(* Logix 5000 project; controller MV vendor 1 type 14 code 217 rev 31.11; software revision 31.00 *)

TASK _1Sec (periodic, rate 1000 ms, priority 10, watchdog 500 ms) : _1Second
TASK MainTask (continuous, watchdog 500 ms) : First_Task, MV_Common, MC_Common, Last_Task

MODULES
   Local : vendor 1 type 14 code 217 (5069 0, rev 31.11)
      FR : vendor 1 type 14 code 217 (Ethernet 192.168.20.32, rev 31.1)
      Remote_IO : vendor 1 type 12 code 298 (Ethernet 192.168.1.1, rev 1.1)
          : vendor 1 type 7 code 76 (Compact 8, rev 1.1, Input RPI 20 ms)
          : vendor 1 type 7 code 76 (Compact 15, rev 1.1, Input RPI 20 ms)
          : 1769-IR6 (Compact 2, rev 1.1, Input RPI 80 ms)
          : 1769-IR6 (Compact 3, rev 1.1, Input RPI 80 ms)
          : 1769-IR6 (Compact 4, rev 1.1, Input RPI 80 ms)
          : 1769-OW16 (Compact 14, rev 1.1, Output RPI 20 ms)
          : vendor 1 type 7 code 79 (Compact 16, rev 3.1, Output RPI 20 ms)
          : 1769-OW16 (Compact 13, rev 1.1, Output RPI 20 ms)
          : 1769-IR6 (Compact 5, rev 1.1, Input RPI 80 ms)
          : vendor 1 type 10 code 47 (Compact 7, rev 1.1, Output RPI 80 ms)
          : 1769-OW16 (Compact 11, rev 1.1, Output RPI 20 ms)
          : vendor 1 type 10 code 47 (Compact 10, rev 1.1, Output RPI 80 ms)
          : 1769-IR6 (Compact 6, rev 1.1, Input RPI 80 ms)
          : 1769-IR6 (Compact 1, rev 1.1, Input RPI 80 ms)
          : vendor 1 type 7 code 79 (Compact 9, rev 3.1, Output RPI 20 ms)
          : 1769-OW16 (Compact 12, rev 1.1, Output RPI 20 ms)
      RIO_Rack_2 : vendor 1 type 12 code 298 (Ethernet 192.168.1.2, rev 1.1)
          : vendor 1 type 7 code 76 (Compact 11, rev 1.1, Input RPI 20 ms)
          : 1769-IQ32 (Compact 14, rev 3.1, Input RPI 20 ms)
          : vendor 1 type 7 code 76 (Compact 4, rev 1.1, Input RPI 20 ms)
          : vendor 1 type 7 code 76 (Compact 7, rev 1.1, Input RPI 20 ms)
          : vendor 1 type 7 code 76 (Compact 6, rev 1.1, Input RPI 20 ms)
          : vendor 1 type 7 code 76 (Compact 12, rev 1.1, Input RPI 20 ms)
          : vendor 1 type 7 code 76 (Compact 9, rev 1.1, Input RPI 20 ms)
          : 1769-IQ32 (Compact 13, rev 3.1, Input RPI 20 ms)
          : vendor 1 type 7 code 79 (Compact 10, rev 3.1, Output RPI 20 ms)
          : vendor 1 type 7 code 79 (Compact 8, rev 3.1, Output RPI 20 ms)
          : vendor 1 type 10 code 48 (Compact 3, rev 1.1, Output RPI 80 ms)
          : 1769-IF4 (Compact 16, rev 3.2, Input RPI 80 ms)
          : vendor 1 type 7 code 73 (Compact 15, rev 3.1, Output RPI 20 ms)
          : vendor 1 type 7 code 79 (Compact 5, rev 3.1, Output RPI 20 ms)
          : 1769-IF8 (Compact 2, rev 1.1, Output RPI 80 ms)
          : 1769-IF8 (Compact 1, rev 1.1, Output RPI 80 ms)
END_MODULES

TYPE CHECKWORD_FLAGS :   // Checkword Flags
STRUCT
   AUTODRV : DINT;   // Auto-Drive Bit No.
   CLOSEDFB : DINT;   // Closed Feedback Bit No.
   OPENFB : DINT;   // Open Feedback Bit No.
   OUTPUT : DINT;   // Output Bit No.
   MANDRV : DINT;   // Manual Drive Bit No.
   MANUAL : DINT;   // Manual Control Bit No.
   CHECKOFF : DINT;   // Checking Off Bit No.
   TRIPPED : DINT;   // Tripped Bit No.
   FAULT : DINT;   // Fault Bit No.
   SIMFAIL : DINT;   // Simulate Failure Bit
   PREVSCAN : DINT;   // Previous Scan State
   FAULTLOGGED : DINT;   // Fault Logged Flag From Scada
   HIGHLIGHT : DINT;   // Highlight on Graphics
   RUNFB : DINT;   // Pump/Drive Run Feedback
   HEALTHYFB : DINT;   // Pump Healthy Feedback
   NOTTRIPPEDFB : DINT;   // Pump Not Tripped Feedback
   HEALTHYFAULTLOGGED : DINT;   // Pump Not Healthy Fault Logged
   TRIPPEDFAULTLOGGED : DINT;   // Pump Tripped Fault Logged
   INPUTSTATUS : DINT;   // Bit Number for Digital Input Status
   INPUTSTATUSDEBOUNCED : DINT;   // Bit Number For Debounced Input Status
   ANALOGSIMULATION : DINT;   // Bit Number For Analog Simulation Enabled
END_STRUCT
END_TYPE

TYPE DateTime :
STRUCT
   Year : DINT;
   Month : DINT;
   Day : DINT;
   Hour : DINT;
   Minute : DINT;
   Second : DINT;
   Microsecond : DINT;
END_STRUCT
END_TYPE

TYPE PlantItem :   // Plant Item
STRUCT
   CW : DINT;   // Checkword
   CheckTime : DINT;   // Check Time
   CheckTimer : DINT;   // Check Time Timer
   DebounceTime : DINT;   // Debounce Time
   DebounceTimer : DINT;   // Debounce Timer
   DriveBits : DINT;   // Item Automatic Drive Bits
   Scaled : REAL;   // Analogue Value Scaled For Input/Output
   RawInput : REAL;   // Raw Input Copied for display On Factory Talk
END_STRUCT
END_TYPE

TYPE Process :   // Data Type For Processes
STRUCT
   Status : DINT;   // Process Current Status
   Step : DINT;   // Process Current Step
   Step_Timer : DINT;   // Current Step Timer
   Fault : DINT;   // Process Current Fault
   Cmd : DINT;   // Command From Scada
   Cmd_avail : DINT;   // Commands Available To Scada
   Cmd_ok : BOOL;   // Startup Command Is Valid Flag
   Cmd_reset : TIMER;   // Startup timer for Invalid Command
   Data_scada : REAL[50];   // Data from Scada
   Data_work : REAL[50];   // Working Data in use by PLC
   Drivebit : DINT;   // Bit Number to Drive Plant Items With
   MessageID : DINT;   // ID to pass with Events/Alarms to Scada
   Past_Prestart : BOOL;   // Flag Set to Indicate past pre start checks.
   Restart_Step : DINT;   // Step to go back to after Continue
END_STRUCT
END_TYPE

TYPE Route :
STRUCT
   CW : DINT;   // Checking Group CW
   CW_Itm : DINT;   // Checking Group Which Has Failed
   Operation : DINT;   // Checking Group Operation Reservation
END_STRUCT
END_TYPE

VAR_GLOBAL   (* controller tags *)
   _1s_pulse : BOOL;
   active : BOOL := 1;
   Alarm_Reset : BOOL;
   alarm_test1 : DINT;
   Always_Off : BOOL;
   Always_On : BOOL := 1;
   Analog_Fault_No : DINT := 30001;
   Analog_Simulation_Enabled : BOOL;
   AT_CUR_PHASE : ALIAS FOR MV_N110[24];   // Phase 0=off 8=Wait yeast 9=Wait Fill 10=Maturation 11to16=Conditioning
   BH_Draindown_ON : DINT;
   CC_CIP_BeerMain_Active : DINT;
   Ch1_cmd_scan_count : DINT;
   Ch1_DataDelay : TIMER := (PRE := 1000);
   Ch2_cmd_scan_count : DINT;
   Ch2_DataDelay : TIMER := (PRE := 1000);
   ChangeDayONS : BOOL;
   CheckTimeMask : INT := 240;
   CIP_AV01_DUMMY_DR : BOOL := 1;
   CIP_AV05_DUMMY_DR : BOOL := 1;
   CIP_AV07_DUMMY_DR : BOOL := 1;
   CIP_AV09_DUMMY_DR : BOOL := 1;
   CLOCK_system_set : BOOL;
   CLOCKsetvalues : DINT[7] := ([0] := 2019, [1] := 3, [2] := 8, [3] := 15, [5] := 1);
        [2]   // Day To Set
        [4]   // Min To Set
        [5]   // Sec to Set
        [0]   // Year To Set
        [3]   // Hour To Set
        [1]   // Month To Set
        [6]   // MS to Set
   colin : DINT := 1237985;
   colon_string : STRING := ':'; {constant}
   comms_to_blunger_write_enabled : BOOL;
   comms_to_fv_route_write_enabled : BOOL;
   comms_to_mv_route_write_enabled : BOOL;
   CurrentTime : DateTime := (Year := 2020, Month := 8, Day := 4, Hour := 17, Second := 6, Microsecond := 778719);
   CWD : CHECKWORD_FLAGS := (CLOSEDFB := 4, OPENFB := 3, OUTPUT := 7, MANDRV := 5, MANUAL := 6, CHECKOFF := 8, FAULT := 15, SIMFAIL := 2, PREVSCAN := 1, FAULTLOGGED := 14, HIGHLIGHT := 9, RUNFB := 3, HEALTHYFB := 10, NOTTRIPPEDFB := 11, HEALTHYFAULTLOGGED := 16, TRIPPEDFAULTLOGGED := 17, INPUTSTATUSDEBOUNCED := 18, ANALOGSIMULATION := 12);
   Default_Check_Time : DINT := 10;
   Delphi_Does_Eng_Func : BOOL;
   Dummy : BOOL := 1;
   enable_comms_to_fv_plc : BOOL := 1;
   Enable_TimeString : BOOL := 1;
   FR_FVS_P01_Consumed : DINT;
   FRHR26_31_Valves_ON_Produced : DINT := 1;
   FT_RT_EMPTYING_SOURCE_VESSEL : DINT;
   FT_RT_FILLING_DESTINATION_VESSEL : DINT;
   FtoF_raw_input : REAL := 5.5534997;
   FV_FLAGS : ALIAS FOR MV_N110[15];   // FLAGS-PROFILE CONTROL
   FV_NUMBER : ALIAS FOR MV_N110[0];   // FV SYSTEM WORKING BUFFER VESSEL NUMBER
   FV_TEMP_BPA : ALIAS FOR MV_N110[1];   // TEMPERATURE BREAKPOINT A. TIME 1/10 HOURS(ALWAYS=0)
   FV_TEMP_BPB : ALIAS FOR MV_N110[3];   // TEMPERATURE BREAKPOINT B. TIME 1/10 HOURS(ALWAYS=0)
   FV_TEMP_BPC : ALIAS FOR MV_N110[5];   // TEMPERATURE BREAKPOINT C. TIME 1/10 HOURS(ALWAYS=0)
   FV_TEMP_BPD : ALIAS FOR MV_N110[7];   // TEMPERATURE BREAKPOINT D. TIME 1/10 HOURS(ALWAYS=0)
   FV_TEMP_BPE : ALIAS FOR MV_N110[9];   // TEMPERATURE BREAKPOINT E. TIME 1/10 HOURS(ALWAYS=0)
   FV_TEMP_BPF : ALIAS FOR MV_N110[11];   // TEMPERATURE BREAKPOINT F. TIME 1/10 HOURS(ALWAYS=0)
   FV_TEMP_BPG : ALIAS FOR MV_N110[13];   // TEMPERATURE BREAKPOINT G. TIME 1/10 HOURS(ALWAYS=0)
   FV_TEMP_SPA : ALIAS FOR MV_N110[2];   // TEMPERATURE SETPOINT A. 1/10 DEGREE 'C'
   FV_TEMP_SPB : ALIAS FOR MV_N110[4];   // TEMPERATURE SETPOINT B. 1/10 DEGREE 'C'
   FV_TEMP_SPC : ALIAS FOR MV_N110[6];   // TEMPERATURE SETPOINT C. 1/10 DEGREE 'C'
   FV_TEMP_SPD : ALIAS FOR MV_N110[8];   // TEMPERATURE SETPOINT D. 1/10 DEGREE 'C'
   FV_TEMP_SPE : ALIAS FOR MV_N110[10];   // TEMPERATURE SETPOINT E. 1/10 DEGREE 'C'
   FV_TEMP_SPF : ALIAS FOR MV_N110[12];   // TEMPERATURE SETPOINT F. 1/10 DEGREE 'C'
   FV_TEMP_SPG : ALIAS FOR MV_N110[14];   // TEMPERATURE SETPOINT G. 1/10 DEGREE 'C'
   FV_YST01_LTX501_AI : PlantItem := (CW := 2#0000_0000_0000_0000_1000_0000_0000_0000, Scaled := 134.09064, RawInput := 18303.0);   // YST01 LTX501
   FV_YST01_LTX501_AI_RawInput : ALIAS FOR RIO_Rack_2:2:I.Ch2Data;
   FV_YST01_LTX501_ALARM : ALARM_DIGITAL;
   FV_YST01_LTX501_Timer_HiLevel : TIMER;
   FV_YST02_LTX501_AI : PlantItem := (CW := 2#0000_0000_0000_0000_1000_0000_0000_0000, Scaled := 140.96251, RawInput := 19036.0);   // YST02 LTX501
   FV_YST02_LTX501_AI_RawInput : ALIAS FOR RIO_Rack_2:2:I.Ch3Data;
   FV_YST02_LTX501_ALARM : ALARM_DIGITAL;
   FV_YST02_LTX501_Timer_HiLevel : TIMER := (PRE := 10000);
   FVHR12_1701 : PlantItem := (CW := 2#0000_0000_0000_0000_0000_0000_0000_1000, CheckTime := 10, CheckTimer := 10);   // Valve FVHR12_17/01
   FVHR12_1701_ALARM : ALARM_DIGITAL;
   FVHR12_1701_CL : ALIAS FOR RIO_Rack_2:13:I.Data.0;   // Valve FVHR12_17/01 Closed
   FVHR12_1701_DR : ALIAS FOR RIO_Rack_2:15:O.Data.0;   // Valve FVHR12_17/01 Drive
   FVHR12_1701_OP : ALIAS FOR RIO_Rack_2:13:I.Data.1;   // Valve FVHR12_17/01 Open
   FVHR12_1702 : PlantItem := (CW := 2#0000_0000_0000_0000_0000_0000_0001_0000, CheckTime := 10, CheckTimer := 10);   // Valve FVHR12_17/02
   FVHR12_1702_ALARM : ALARM_DIGITAL;
   FVHR12_1702_CL : ALIAS FOR RIO_Rack_2:13:I.Data.2;   // Valve FVHR12_17/02 Closed
   FVHR12_1702_DR : ALIAS FOR RIO_Rack_2:15:O.Data.1;   // Valve FVHR12_17/02 Drive
   FVHR12_1702_OP : ALIAS FOR RIO_Rack_2:13:I.Data.3;   // Valve FVHR12_17/02 Open
   FVHR12_1703 : PlantItem := (CW := 2#0000_0000_0000_0000_0000_0000_0001_0000, CheckTime := 10, CheckTimer := 10);   // Valve FVHR12_17/03
   FVHR12_1703_ALARM : ALARM_DIGITAL;
   FVHR12_1703_CL : ALIAS FOR RIO_Rack_2:13:I.Data.10;   // Valve FVHR12_17/03 Closed
   FVHR12_1703_DR : ALIAS FOR RIO_Rack_2:15:O.Data.5;   // Valve FVHR12_17/03 Drive
   FVHR12_1703_OP : ALIAS FOR RIO_Rack_2:13:I.Data.11;   // Valve FVHR12_17/03 Open
   FVHR12_17_Valves_ON : BOOL := 1;   // Check bit to confirm valves for FV12-17 route are open
   FVHR18_21_Valves_ON : BOOL := 1;   // Check bit to confirm valves for FV18-21 route are open
   FVHR18_2501 : PlantItem := (CW := 2#0000_0000_0000_0000_0000_0000_0000_1000, CheckTime := 10, CheckTimer := 10);   // Valve FVHR18_25/01
   FVHR18_2501_ALARM : ALARM_DIGITAL;
   FVHR18_2501_CL : ALIAS FOR RIO_Rack_2:13:I.Data.18;   // Valve FVHR18_25/01 Closed
   FVHR18_2501_DR : ALIAS FOR RIO_Rack_2:15:O.Data.9;   // Valve FVHR18_25/01 Drive
   FVHR18_2501_OP : ALIAS FOR RIO_Rack_2:13:I.Data.19;   // Valve FVHR18_25/01 Open
   FVHR18_2502 : PlantItem := (CW := 2#0000_0000_0000_0000_0000_0000_0001_0000, CheckTime := 10, CheckTimer := 10);   // Valve FVHR18_25/02
   FVHR18_2502_ALARM : ALARM_DIGITAL;
   FVHR18_2502_CL : ALIAS FOR RIO_Rack_2:13:I.Data.20;   // Valve FVHR18_25/02 Closed
   FVHR18_2502_DR : ALIAS FOR RIO_Rack_2:15:O.Data.10;   // Valve FVHR18_25/02 Drive
   FVHR18_2502_OP : ALIAS FOR RIO_Rack_2:13:I.Data.21;   // Valve FVHR18_25/02 Open
   FVHR18_2503 : PlantItem := (CW := 2#0000_0000_0000_0000_0000_0000_0000_1000, CheckTime := 10, CheckTimer := 10);   // Valve FVHR18_25/03
   FVHR18_2503_ALARM : ALARM_DIGITAL;
   FVHR18_2503_CL : ALIAS FOR RIO_Rack_2:13:I.Data.22;   // Valve FVHR18_25/03 Closed
   FVHR18_2503_DR : ALIAS FOR RIO_Rack_2:15:O.Data.11;   // Valve FVHR18_25/03 Drive
   FVHR18_2503_OP : ALIAS FOR RIO_Rack_2:13:I.Data.23;   // Valve FVHR18_25/03 Open
   FVHR18_2504 : PlantItem := (CW := 2#0000_0000_0000_0000_0000_0000_0001_0000, CheckTime := 10, CheckTimer := 10);   // Valve FVHR18_25/04
   FVHR18_2504_ALARM : ALARM_DIGITAL;
   FVHR18_2504_CL : ALIAS FOR RIO_Rack_2:13:I.Data.24;   // Valve FVHR18_25/04 Closed
   FVHR18_2504_DR : ALIAS FOR RIO_Rack_2:15:O.Data.12;   // Valve FVHR18_25/04 Drive
   FVHR18_2504_OP : ALIAS FOR RIO_Rack_2:13:I.Data.25;   // Valve FVHR18_25/04 Open
   FVHR18_2505 : PlantItem := (CW := 2#0000_0000_0000_0000_0000_0000_0001_0000, CheckTime := 10, CheckTimer := 10);   // Valve FVHR18_25/05
   FVHR18_2505_ALARM : ALARM_DIGITAL;
   FVHR18_2505_CL : ALIAS FOR RIO_Rack_2:13:I.Data.26;   // Valve FVHR18_25/05 Closed
   FVHR18_2505_DR : ALIAS FOR RIO_Rack_2:15:O.Data.13;   // Valve FVHR18_25/05 Drive
   FVHR18_2505_OP : ALIAS FOR RIO_Rack_2:13:I.Data.27;   // Valve FVHR18_25/05 Open
   FVHR18_2506 : PlantItem := (CW := 2#0000_0000_0000_0000_0000_0000_0001_0000, CheckTime := 10, CheckTimer := 10);   // Valve FVHR18_25/06
   FVHR18_2506_ALARM : ALARM_DIGITAL;
   FVHR18_2506_CL : ALIAS FOR RIO_Rack_2:13:I.Data.28;   // Valve FVHR18_25/06 Closed
   FVHR18_2506_DR : ALIAS FOR RIO_Rack_2:15:O.Data.14;   // Valve FVHR18_25/06 Drive
   FVHR18_2506_OP : ALIAS FOR RIO_Rack_2:13:I.Data.29;   // Valve FVHR18_25/06 Open
   FVHR1_1101 : PlantItem := (CW := 2#0000_0000_0000_0000_0000_0000_0000_1000, CheckTime := 10, CheckTimer := 10);   // Valve FVHR1_11/01
   FVHR1_1101_ALARM : ALARM_DIGITAL;
   FVHR1_1101_CL : ALIAS FOR RIO_Rack_2:13:I.Data.4;   // Valve FVHR1_11/01 Closed
   FVHR1_1101_DR : ALIAS FOR RIO_Rack_2:15:O.Data.2;   // Valve FVHR1_11/01 Drive
   FVHR1_1101_OP : ALIAS FOR RIO_Rack_2:13:I.Data.5;   // Valve FVHR1_11/01 Open
   FVHR1_1102 : PlantItem := (CW := 2#0000_0000_0000_0000_0000_0000_0001_0000, CheckTime := 10, CheckTimer := 10);   // Valve FVHR1_11/02
   FVHR1_1102_ALARM : ALARM_DIGITAL;
   FVHR1_1102_CL : ALIAS FOR RIO_Rack_2:13:I.Data.6;   // Valve FVHR1_11/02 Closed
   FVHR1_1102_DR : ALIAS FOR RIO_Rack_2:15:O.Data.3;   // Valve FVHR1_11/02 Drive
   FVHR1_1102_OP : ALIAS FOR RIO_Rack_2:13:I.Data.7;   // Valve FVHR1_11/02 Open
   FVHR1_1103 : PlantItem := (CW := 2#0000_0000_0000_0000_0000_0000_0001_0000, CheckTime := 10, CheckTimer := 10);   // Valve FVHR1_11/03
   FVHR1_1103_ALARM : ALARM_DIGITAL;
   FVHR1_1103_CL : ALIAS FOR RIO_Rack_2:13:I.Data.8;   // Valve FVHR1_11/03 Closed
   FVHR1_1103_DR : ALIAS FOR RIO_Rack_2:15:O.Data.4;   // Valve FVHR1_11/03 Drive
   FVHR1_1103_OP : ALIAS FOR RIO_Rack_2:13:I.Data.9;   // Valve FVHR1_11/03 Open
   FVHR1_11_Valves_ON : BOOL := 1;   // Check bit to confirm valves for FV1-11 route are open
   FVHR1_1701 : PlantItem := (CW := 2#0000_0000_0000_0000_0000_0000_0001_0000, CheckTime := 10, CheckTimer := 10);   // Valve FVHR1_17/01
   FVHR1_1701_ALARM : ALARM_DIGITAL;
   FVHR1_1701_CL : ALIAS FOR RIO_Rack_2:13:I.Data.16;   // Valve FVHR1_17/01 Closed
   FVHR1_1701_DR : ALIAS FOR RIO_Rack_2:15:O.Data.8;   // Valve FVHR1_17/01 Drive
   FVHR1_1701_OP : ALIAS FOR RIO_Rack_2:13:I.Data.17;   // Valve FVHR1_17/01 Open
   FVHR22_25_Valves_ON : BOOL := 1;   // Check bit to confirm valves for FV22-25 route are open
   FVHR26_3101 : PlantItem := (CW := 2#0000_0000_0000_0000_0000_0000_0000_1000, CheckTime := 10, CheckTimer := 10);   // Valve FVHR26_31/01
   FVHR26_3101_ALARM : ALARM_DIGITAL;
   FVHR26_3101_CL : ALIAS FOR RIO_Rack_2:14:I.Data.2;   // Valve FVHR26_31/01 Closed
   FVHR26_3101_DR : ALIAS FOR RIO_Rack_2:15:O.Data.17;   // Valve FVHR26_31/01 Drive
   FVHR26_3101_OP : ALIAS FOR RIO_Rack_2:14:I.Data.3;   // Valve FVHR26_31/01 Open
   FVHR26_3102 : PlantItem := (CW := 2#0000_0000_0000_0000_0000_0000_0001_0000, CheckTime := 10, CheckTimer := 10);   // Valve FVHR26_31/02
   FVHR26_3102_ALARM : ALARM_DIGITAL;
   FVHR26_3102_CL : ALIAS FOR RIO_Rack_2:14:I.Data.4;   // Valve FVHR26_31/02 Closed
   FVHR26_3102_DR : ALIAS FOR RIO_Rack_2:15:O.Data.18;   // Valve FVHR26_31/02 Drive
   FVHR26_3102_OP : ALIAS FOR RIO_Rack_2:14:I.Data.5;   // Valve FVHR26_31/02 Open
   FVHR26_3103 : PlantItem := (CW := 2#0000_0000_0000_0000_0000_0000_0001_0000, CheckTime := 10, CheckTimer := 10);   // Valve FVHR26_31/03
   FVHR26_3103_ALARM : ALARM_DIGITAL;
   FVHR26_3103_CL : ALIAS FOR RIO_Rack_2:14:I.Data.6;   // Valve FVHR26_31/03 Closed
   FVHR26_3103_DR : ALIAS FOR RIO_Rack_2:15:O.Data.19;   // Valve FVHR26_31/03 Drive
   FVHR26_3103_OP : ALIAS FOR RIO_Rack_2:14:I.Data.7;   // Valve FVHR26_31/03 Open
   FVHR26_31_Valves_ON : BOOL := 1;   // Check bit to confirm valves for FV26-31 route are open
   FVHRCH201 : PlantItem := (CW := 2#0000_0000_0000_0000_0000_0000_0001_0000, CheckTime := 10, CheckTimer := 10);   // Valve FVHRCH201
   FVHRCH201_ALARM : ALARM_DIGITAL;
   FVHRCH201_CL : ALIAS FOR RIO_Rack_2:14:I.Data.10;   // Valve FVHRCH201 Closed
   FVHRCH201_DR : ALIAS FOR RIO_Rack_2:15:O.Data.21;   // Valve FVHRCH201 Drive
   FVHRCH201_OP : ALIAS FOR RIO_Rack_2:14:I.Data.11;   // Valve FVHRCH201 Open
   FVHRCH202 : PlantItem := (CW := 2#0000_0000_0000_0000_0000_0000_0001_0000, CheckTime := 10, CheckTimer := 10);   // Valve FVHRCH202
   FVHRCH202_ALARM : ALARM_DIGITAL;
   FVHRCH202_CL : ALIAS FOR RIO_Rack_2:14:I.Data.14;   // Valve FVHRCH202 Closed
   FVHRCH202_DR : ALIAS FOR RIO_Rack_2:15:O.Data.23;   // Valve FVHRCH202 Drive
   FVHRCH202_OP : ALIAS FOR RIO_Rack_2:14:I.Data.15;   // Valve FVHRCH202 Open
   FVHRCW01 : PlantItem := (CW := 2#0000_0000_0000_0000_0000_0000_0001_0000, CheckTime := 10, CheckTimer := 10);   // Valve FVHRCW01
   FVHRCW01_ALARM : ALARM_DIGITAL;
   FVHRCW01_CL : ALIAS FOR RIO_Rack_2:14:I.Data.12;   // Valve FVHRCW01 Closed
   FVHRCW01_DR : ALIAS FOR RIO_Rack_2:15:O.Data.22;   // Valve FVHRCW01 Drive
   FVHRCW01_OP : ALIAS FOR RIO_Rack_2:14:I.Data.13;   // Valve FVHRCW01 Open
   FVHRFM03_ALARM : ALARM_DIGITAL;
   FVHRFM03_IP : PlantItem := (CW := 2#0000_0000_0000_0000_1000_0000_0000_0000, CheckTime := 15, CheckTimer := 15, Scaled := -0.1125, RawInput := 3996.0);   // Flow Meter Transmitter
   FVHRFM03_IP_RawInput : ALIAS FOR RIO_Rack_2:16:I.Ch2Data;   // Flow Meter Raw Data
   FVHRLTX02_ALARM : ALARM_DIGITAL;
   FVHRLTX02_IP : PlantItem := (CW := 2#0000_0000_0000_0000_1000_0000_0000_0000, CheckTime := 15, CheckTimer := 15, Scaled := 307.71875, RawInput := 13847.0);   // Effluent Tank Level Transmitter
   FVHRLTX02_IP_Percentage : DINT := 62;
   FVHRLTX02_IP_RawInput : ALIAS FOR RIO_Rack_2:16:I.Ch1Data;   // Effluent Tank Level Transmitter Raw Data
   FVHRLTX02_Timer_HiLevel : TIMER := (PRE := 10000);
   FVHRM01 : PlantItem := (CW := 2#0000_0000_0000_0000_0000_0000_0001_0000, CheckTime := 10, CheckTimer := 10);   // Valve FVHRM01
   FVHRM01_ALARM : ALARM_DIGITAL;
   FVHRM01_CL : ALIAS FOR RIO_Rack_2:13:I.Data.30;   // Valve FVHRM01 Closed
   FVHRM01_DR : ALIAS FOR RIO_Rack_2:15:O.Data.15;   // Valve FVHRM01 Drive
   FVHRM01_OP : ALIAS FOR RIO_Rack_2:13:I.Data.31;   // Valve FVHRM01 Open
   FVHRM02 : PlantItem := (CW := 2#0000_0000_0000_0000_0000_0000_0001_0000, CheckTime := 10, CheckTimer := 10);   // Valve FVHRM02
   FVHRM02_ALARM : ALARM_DIGITAL;
   FVHRM02_CL : ALIAS FOR RIO_Rack_2:14:I.Data.0;   // Valve FVHRM02 Closed
   FVHRM02_DR : ALIAS FOR RIO_Rack_2:15:O.Data.16;   // Valve FVHRM02 Drive
   FVHRM02_OP : ALIAS FOR RIO_Rack_2:14:I.Data.1;   // Valve FVHRM02 Open
   FVHRM03 : PlantItem := (CW := 2#0000_0000_0000_0000_0000_0000_0001_0000, CheckTime := 10, CheckTimer := 10);   // Valve FVHRM03
   FVHRM03_ALARM : ALARM_DIGITAL;
   FVHRM03_CL : ALIAS FOR RIO_Rack_2:14:I.Data.8;   // Valve FVHRM03 Closed
   FVHRM03_DR : ALIAS FOR RIO_Rack_2:15:O.Data.20;   // Valve FVHRM03 Drive
   FVHRM03_OP : ALIAS FOR RIO_Rack_2:14:I.Data.9;   // Valve FVHRM03 Open
   FVHRM04 : PlantItem := (CW := 2#0000_0000_0000_0000_0000_0000_0001_0000, CheckTime := 10, CheckTimer := 10);   // Valve FVHRM04
   FVHRM04_ALARM : ALARM_DIGITAL;
   FVHRM04_CL : ALIAS FOR RIO_Rack_2:13:I.Data.12;   // Valve FVHRM04 Closed
   FVHRM04_DR : ALIAS FOR RIO_Rack_2:15:O.Data.6;   // Valve FVHRM04 Drive
   FVHRM04_OP : ALIAS FOR RIO_Rack_2:13:I.Data.13;   // Valve FVHRM04 Open
   FVHRMD01 : PlantItem := (CW := 2#0000_0000_0000_0000_0000_0000_0000_1000, CheckTime := 10, CheckTimer := 10);   // Valve FVHRMD01
   FVHRMD01_ALARM : ALARM_DIGITAL;
   FVHRMD01_CL : ALIAS FOR RIO_Rack_2:13:I.Data.14;   // Valve FVHRMD01 Closed
   FVHRMD01_DR : ALIAS FOR RIO_Rack_2:15:O.Data.7;   // Valve FVHRMD01 Drive
   FVHRMD01_OP : ALIAS FOR RIO_Rack_2:13:I.Data.15;   // Valve FVHRMD01 Open
   FVHRTM01_ALARM : ALIAS FOR RIO_Rack_2:14:I.Data.16;   // Turbidty Meter FVHRTM01 Fault
   FVHRTM01_IP : PlantItem := (CW := 2#0000_0000_0000_0000_1000_0000_0000_0000, CheckTime := 15, CheckTimer := 15, Scaled := 0.012496876, RawInput := 3998.0);   // Turbidty Meter FVHRTM01
   FVHRTM01_IP_RawInput : ALIAS FOR RIO_Rack_2:16:I.Ch0Data;   // Turbidty Meter FVHRTM01 Raw Data
   fvrroute_slc_still_active : BOOL;
   Half_Second_Timer_Off : TIMER;
   Half_Second_Timer_On : TIMER := (PRE := 1000, ACC := 644, EN := 1, TT := 1);
   Half_Second_Toggle : BOOL;
   hr_string : STRING := '0';
   IGI_TestBit : BOOL := 1;
   indirect_bit_temp : INT := 42;
   Item_Faults_Are_Latched : BOOL;
   Item_Simulation_Flag : BOOL;
   ItoF_raw_input : INT := 3945;
   MC_ALARM_RETURNED_STRING : STRING := 'CH1_R1 feedbacks have failed.';
   MC_B12 : INT[255] := ([0] := -3698, [1] := -29, [2] := -513);   // PX SWITCH Proxy switch flags f ile
        [1].2   // Prog 18: Centr.beer main + CT transfer p/x switches ok
        [1].4   // Prog.20: Yeast Suction Main FVs 18-25 Short p/x switches ok
        [2].2   // Prog.34: Yeast Suction Main FVs 26-31 Short p/x switches ok
        [2].5   // Prog 37: Yeast Suction Main FVs 1-17 Long p/x switches ok
        [2].6   // Prog 38: Yeast Suction Main FVs 18- 25 Long p/x switches ok
        [1].13   // Prog.29: MVs 36-47 filling main p/x switches ok
        [2].7   // Prog 39: Yeast Suction Main FVs 26- 31 Long p/x switches ok
        [0].11   // Prog.11: Centr.beer main only p/x switches ok
        [0].13   // Prog.13: MVs 3-4/ 8-10/23/YPV p/x switches ok
        [1].5   // Prog.21: Yeast Room Main + Pump p/x switches ok
        [0].14   // Prog.14: MVs 30-35/ YSV3 p/x switches ok
        [1].0   // Prog.16: MVs 11-13/ 17-19 p/x switches ok
        [1].3   // Prog.19: Yeast Suction Main FVs 1-17 Short p/x switches ok
        [2].8   // Prog 40: PVPP Mixing Tank p/x switches ok
        [2].0   // Prog.32: MVs 36-47 racking main 3 p/x switches ok
        [0].8   // Prog.8: Yeast suction main p/x switches ok
        [2].10   // Prog.42: Gales Yeast Main p/x switches ok
        [0].4   // Prog.4: YSV 1 p/x switches ok
        [0].5   // Prog.5: YSV 2 p/x switches ok
        [1].6   // Prog 22: YCV1 p/x switches ok
        [1].7   // Prog 23: YCV2 p/x switches ok
        [1].8   // Prog 24: YCV3 p/x switches ok
        [3].0   // Prog.48: FV Bypass Line switches ok
        [0].15   // Prog.15: MVs 14-16/ 20-22 p/x switches ok
        [0].6   // Prog.6: YSV1 reseeding line p/x switches ok
        [0].7   // Prog.7: Yeast pitching main p/x switches ok
        [0].12   // Prog.12 MVs 1-2/5-7 p/x switches ok
        [0].10   // Prog.10: Centrifuges p/x switches ok
        [1].10   // Prog.26: WYSTs 1 & 2 p/x switches ok
        [0].1   // Prog.1: FVs 1-17 p/x switches ok
        [1].9   // Prog.25: Filtrate Tank p/x switches ok
        [2].3   // Prog.35: Filtrate main p/x switches ok
        [1].1   // Prog.17: Racking main p/x switches ok
        [1].11   // Prog.27: MVs 36-47 p/x switches ok
        [1].12   // Prog.28: FVs 26-31 p/x switches ok
        [1].14   // Prog.30: MVs 36-47 racking main 1 p/x switches ok
        [2].4   // Prog.36: Yeast Press p/x switches ok
        [1].15   // Prog.31: MVs 36-47 racking main 2 p/x switches ok
        [2].1   // Prog.33: FVs 26-31 green beer mains p/x switches ok
        [2].9   // Prog.41: Gales Green Beer Main p/x switches ok
        [0].9   // Prog.9: Green beer main p/x switches ok
        [0].2   // Prog.2: FVs 18-21 p/x switches ok
        [0].3   // Prog.3: FVs 22-25 p/x switches ok
   MC_B240 : INT[255];   // CH1 RN PMP Channel 1 return pum p drive flags
        [1].0   // CH1 drive prog.no.16 return pump flag
        [1].3   // CH1 drive prog.no.19 return pump flag
        [1].6   // CH1 drive prog no.22 return pump flag
        [1].7   // CH1 drive prog no.23 return pump flag
        [1].8   // CH1 drive prog no.24 return pump flag
        [1].9   // CH1 drive prog no.25 return pump flag
        [0].1   // CH1 drive prog.no.1 return pump flag
        [0].2   // CH1 drive prog.no.2 return pump flag
        [0].3   // CH1 drive prog.no.3 return pump flag
        [0].4   // CH1 drive prog.no.4 return pump flag
        [0].5   // CH1 drive prog.no.5 return pump flag
        [0].6   // CH1 drive prog.no.6 return pump flag
        [0].8   // CH1 drive prog.no.8 return pump flag
        [0].12   // CH1 drive prog.no.12 return pump flag
        [0].13   // CH1 drive prog.no.13 return pump flag
        [0].14   // CH1 drive prog.no.14 return pump flag
        [0].15   // CH1 drive prog.no.15 return pump flag
        [1].10   // CH1 drive prog no.26 return pump flag
   MC_B241 : INT[255];   // CH2 RN PMP Channel 2 return pum p drive flags
        [1].0   // CH2 drive prog.no.16 return pump flag
        [1].3   // CH2 drive prog.no.19 return pump flag
        [1].6   // CH2 drive prog no.22 return pump flag
        [1].7   // CH2 drive prog no.23 return pump flag
        [1].8   // CH2 drive prog no.24 return pump flag
        [1].9   // CH2 drive prog no.25 return pump flag
        [0].1   // CH2 drive prog.no.1 return pump flag
        [0].2   // CH2 drive prog.no.2 return pump flag
        [0].3   // CH2 drive prog.no.3 return pump flag
        [0].4   // CH2 drive prog.no.4 return pump flag
        [0].5   // CH2 drive prog.no.5 return pump flag
        [0].6   // CH2 drive prog.no.6 return pump flag
        [0].8   // CH2 drive prog.no.8 return pump flag
        [0].12   // CH2 drive prog.no.12 return pump flag
        [0].13   // CH2 drive prog.no.13 return pump flag
        [0].14   // CH1 drive prog.no.14 return pump flag
        [0].15   // CH2 drive prog.no.15 return pump flag
        [1].10   // CH2 drive prog no.26 return pump flag
   MC_B242 : INT[255] := ([1] := 2);   // CH1 ROUTE Channel 1 route requ est flags
        [1].0   // CH1 drive prog.no.16 routing valves
        [1].2   // CH1 drive prog.no.18 routing valves
        [1].3   // CH1 drive prog.no.19 routing valves
        [1].4   // CH1 drive prog.no.20 routing valves
        [1].5   // CH1 drive prog.no.21 routing valves
        [0].12   // CH1 drive prog.no.12 routing valves
        [0].13   // CH1 drive prog.no.13 routing valves
        [0].14   // CH1 drive prog.no.14 routing valves
        [0].15   // CH1 drive prog.no.15 routing valves
        [2].10   // CH1 drive prog.no.42 routing valves
   MC_B243 : INT[255];   // CH2 ROUTE Channel 2 route requ est flags
        [1].0   // CH2 drive prog.no.16 routing valves
        [1].2   // CH2 drive prog.no.18 routing valves
        [1].3   // CH2 drive prog.no.19 routing valves
        [1].4   // CH2 drive prog.no.20 routing valves
        [1].5   // CH2 drive prog.no.21 routing valves
        [0].12   // CH2 drive prog.no.12 routing valves
        [0].13   // CH2 drive prog.no.13 routing valves
        [0].14   // CH2 drive prog.no.14 routing valves
        [0].15   // CH2 drive prog.no.15 routing valves
        [2].10   // CH2 drive prog.no 42 routing valves
   MC_B3 : INT[255];   // BINARY
        [0].0   // *********** Simulation Enabled ***********
        [0].1   // Time/Date Setting oneshot
        [0].2   // Settings reload oneshot
   MC_B3_0_1_OUTPUTBIT : BOOL;
   MC_B3_0_2_OUTPUTBIT : BOOL;
   MC_bit_data_file_address : DINT := 243;
   MC_bit_file_bit_offset : DINT;
   MC_bit_file_word_offset : DINT;
   MC_bit_offset : DINT := 17;
   MC_bit_returned : BOOL := 1;
   MC_bit_value_to_set : DINT;
   MC_CD_T1 : PlantItem := (CW := 2#0000_0000_0000_0000_0000_0000_0001_0000, CheckTime := 8, CheckTimer := 8);   // CD_T1
   MC_CD_T1_ALARM : ALARM_DIGITAL;
   MC_CD_T1_C : ALIAS FOR RIO_Rack_2:7:I.Data.23;
   MC_CD_T1_DR : ALIAS FOR RIO_Rack_2:8:O.Data.11;
   MC_CD_T1_O : ALIAS FOR RIO_Rack_2:7:I.Data.19;
   MC_CD_T2 : PlantItem := (CW := 2#0000_0000_0000_0000_0000_0000_0001_0000, CheckTime := 8, CheckTimer := 8);   // CD_T2
   MC_CD_T2_ALARM : ALARM_DIGITAL;
   MC_CD_T2_C : ALIAS FOR RIO_Rack_2:7:I.Data.28;
   MC_CD_T2_DR : ALIAS FOR RIO_Rack_2:8:O.Data.12;
   MC_CD_T2_O : ALIAS FOR RIO_Rack_2:7:I.Data.24;
   MC_CH1_ACTIVE : ALIAS FOR MC_N100[30].1;   // CH1 active flag
   MC_CH1_CIP_Messages : STRING[20] := ([0] := 'Racking Main Normal clean', [1] := 'Detergent 1 of 1', [2] := '00:01:25', [3] := '00:16:25', [5] := '17:07:10');   // CH1 CIP Scada Messages
        [5]   // Channel 1 CIP Completion Clock Time
        [3]   // Channel 1 CIP Total Time Text for Scada
        [1]   // Channel 1 CIP Cycle Text for Scada
        [0]   // Channel 1 CIP Program Text for Scada
        [2]   // Channel 1 CIP Time Left Text for Scada
        [4]   // Channel 1 CIP Down Time Text for Scada
   MC_CH1_CIP_Misc : DINT[20] := ([0] := 1409, [1] := 425);
   MC_CH1_CIP_MiscReal : REAL[20] := ([0] := 30.092262);
   MC_CH1_CSTEP : ALIAS FOR MC_N100[34];   // CH1 command processor current step
   MC_CH1_CTX1_AI : PlantItem := (CW := 2#0000_0000_0000_0000_1000_0000_0000_0000, CheckTime := 15, CheckTimer := 15, Scaled := 2.73125, RawInput := 8370.0);   // CH1_CTX1
   MC_CH1_CTX1_AI_RawInput : ALIAS FOR RIO_Rack_2:1:I.Ch2Data;   // Real Analog Input , Do Not Use In Code
   MC_CH1_CYCDONE : ALIAS FOR MC_T105[2].DN;   // CH1 current cycle complete
   MC_CH1_CYCLE : ALIAS FOR MC_N100[1];   // CH1 current CIP cycle
   MC_CH1_Delay_For_Data : TIMER := (PRE := 2000);
   MC_CH1_DETRTN : ALIAS FOR MC_N100[18].1;   // CH1 Is Detergent Return flag
   MC_CH1_DONE : ALIAS FOR MC_N100[30].4;   // CH1 cycle complete flag
   MC_CH1_DR1 : PlantItem := (CW := 2#0000_0000_0000_0000_0000_0000_1000_1011, CheckTime := 20, CheckTimer := 20, DriveBits := 1);   // CH1_DR1
   MC_CH1_DR1_ALARM : ALARM_DIGITAL;
   MC_CH1_DR1_C : ALIAS FOR RIO_Rack_2:4:I.Data.30;
   MC_CH1_DR1_DR : ALIAS FOR RIO_Rack_2:5:O.Data.14;
   MC_CH1_DR1_O : ALIAS FOR RIO_Rack_2:4:I.Data.26;
   MC_CH1_DR2 : PlantItem := (CW := 2#0000_0000_0000_0000_0000_0000_0001_0000, CheckTime := 8, CheckTimer := 8);   // CH1_DR2
   MC_CH1_DR2_ALARM : ALARM_DIGITAL;
   MC_CH1_DR2_C : ALIAS FOR RIO_Rack_2:4:I.Data.31;
   MC_CH1_DR2_DR : ALIAS FOR RIO_Rack_2:5:O.Data.15;
   MC_CH1_DR2_O : ALIAS FOR RIO_Rack_2:4:I.Data.27;
   MC_CH1_DRAIN : PlantItem := (CW := 2#0000_0000_0000_0000_0000_0000_0001_0000, CheckTime := 20, CheckTimer := 20);   // CH1_DRAIN
   MC_CH1_DRAIN_ALARM : ALARM_DIGITAL;
   MC_CH1_DRAIN_C : ALIAS FOR RIO_Rack_2:4:I.Data.28;
   MC_CH1_DRAIN_DR : ALIAS FOR RIO_Rack_2:5:O.Data.12;
   MC_CH1_DRAIN_O : ALIAS FOR RIO_Rack_2:4:I.Data.24;
   MC_CH1_DT : ALIAS FOR MC_N100[10];   // CH1 detergent tank to use (1 or 2)
   MC_CH1_DT1 : PlantItem := (CW := 2#0000_0000_0000_0000_0000_0000_1000_1011, CheckTime := 8, CheckTimer := 8, DriveBits := 1);   // CH1_DT1
   MC_CH1_DT1_ALARM : ALARM_DIGITAL;
   MC_CH1_DT1_C : ALIAS FOR RIO_Rack_2:6:I.Data.4;
   MC_CH1_DT1_DR : ALIAS FOR RIO_Rack_2:5:O.Data.16;
   MC_CH1_DT1_O : ALIAS FOR RIO_Rack_2:6:I.Data.0;
   MC_CH1_DT2 : PlantItem := (CW := 2#0000_0000_0000_0000_0000_0000_0001_0000, CheckTime := 8, CheckTimer := 8);   // CH1_DT2
   MC_CH1_DT2_ALARM : ALARM_DIGITAL;
   MC_CH1_DT2_C : ALIAS FOR RIO_Rack_2:6:I.Data.5;
   MC_CH1_DT2_DR : ALIAS FOR RIO_Rack_2:5:O.Data.17;
   MC_CH1_DT2_O : ALIAS FOR RIO_Rack_2:6:I.Data.1;
   MC_CH1_EVENT : ALIAS FOR MC_N100[23];   // CH1 event register
   MC_CH1_EXTEND : ALIAS FOR MC_N100[30].5;   // CH1 extend cycle flag
   MC_CH1_FAULT : ALIAS FOR MC_N100[20];   // CH1 fault register
   MC_CH1_FM_AI : PlantItem := (CW := 2#0000_0000_0000_0000_1000_0000_0000_0000, CheckTime := 15, CheckTimer := 15, Scaled := 199.3125, RawInput := 10378.0);   // CH1_FM
   MC_CH1_FM_AI_RawInput : ALIAS FOR RIO_Rack_2:1:I.Ch4Data;   // Real Analog Input , Do Not Use In Code
   MC_CH1_ISLINE : ALIAS FOR MC_N102[13].0;   // CH1 Is Line Clean flag
   MC_CH1_LF1 : PlantItem := (CW := 2#0000_0000_0000_0000_0000_0001_0001_0000, CheckTime := 8, CheckTimer := 8);   // CH1_LF1
   MC_CH1_LF1_ALARM : ALARM_DIGITAL;
   MC_CH1_LF1_C : ALIAS FOR RIO_Rack_2:6:I.Data.7;
   MC_CH1_LF1_DR : ALIAS FOR RIO_Rack_2:5:O.Data.19;
   MC_CH1_LF1_O : ALIAS FOR RIO_Rack_2:6:I.Data.3;